// TIA Portal project "e045002v089" (V13) (continued)
VAR_GLOBAL   // PLC tag table "I/O Intercambio Envolvedora"
   "iPalletRetractil" AT %E2.0 : Bool;   // Pallet retractilado (desde el retractilador)
   "oRetractiSeg" AT %A17.7 : Bool;   // Retractilador Seguridades (hacia Retractilador)
   "iPeticionPallet" AT %E2.1 : Bool;   // Petición de pallet (desde el retractilador)
   "oRetractiPermiso" AT %A17.6 : Bool;   // Retractilador Permiso (hacia Retractilador)
   "iBrazoPos_Envolv" AT %E10.5 : Bool;   // Brazo en posición y Freno cerrado en Envolvedora (Retractilador)
   "oHabilMovBrazo_Envol" AT %A16.3 : Bool;   // Habilitación apertura freno brazo Envolvedora (Retractilador)
END_VAR

VAR_GLOBAL   // PLC tag table "I/O Intercambio Cartonero"
   "iCartZonaSeg" AT %M230.1 : Bool;   // Señal de Cartonero: 1= Fuera de zona de paletizadora
   "iCartAplicado" AT %M230.2 : Bool;   // Señal de Cartonero: 1= Cartón aplicado
   "oTomarCartón" AT %A34.3 : Bool;   // Señal a Cartonero: 1= Tomar cartón
   "oAplicarCartón" AT %A34.4 : Bool;   // Señal a Cartonero: 1= Aplicar Cartón
   "oPaleZonaSeg" AT %A34.5 : Bool;   // Señal a Cartonero: 1= Paletizadora en zona segura para el cartonero
   "oPaleSinAlarm" AT %A34.6 : Bool;   // Señal a Cartonero: 1= Paletizadora sin alarmas
   "iCartSinAlarm" AT %M230.0 : Bool;   // Señal de Cartonero: 1= Sin Alarmas
END_VAR

VAR_GLOBAL   // PLC tag table "260_EtiquetadoraYFechadoras"
   "i_FallEnEtiq" AT %I6.6 : Bool;
   "i_FallEnFechadora1" AT %I10.6 : Bool;
   "iSns_PresCajaEmpujador" AT %I11.0 : Bool;
END_VAR

TYPE "Filas_Receta"
   STRUCT
      Bit_1_Elemento : Array [1..10] of Bool;
      Bit_2_Elemento : Array [1..10] of Bool;
   END_STRUCT;
END_TYPE

TYPE "Capas_Receta"
   STRUCT
      Filas : Array [1..6] of "Filas_Receta";
      Usar_Pistón : Bool;
   END_STRUCT;
END_TYPE

TYPE "Elementos HMI"
   STRUCT
      Figura : Byte;
      Estado : Byte;
      Offset_X : Int;
   END_STRUCT;
END_TYPE

TYPE "Filas HMI"
   STRUCT
      Offset_Y : Int;
      Elemento : Array [1 .. 10] of "Elementos HMI";
   END_STRUCT;
END_TYPE

TYPE "Filas_Proceso"
   STRUCT
      Bit_1_Elemento : Array [1 .. 10] of Bool;
      Bit_2_Elemento : Array [1 .. 10] of Bool;
      Actual_Elemento : Array [1 .. 10] of Bool;
   END_STRUCT;
END_TYPE

TYPE "Capas_Proceso"
   STRUCT
      Fila : Array [1 .. 6] of "Filas_Proceso";
      Usar_Pistón : Bool;
   END_STRUCT;
END_TYPE

TYPE "PETICION_CONTROL"
   STRUCT
      cero : Byte;
      PETICION : Byte;
      PARAMETRO : Array [1 .. 3] of Word;
   END_STRUCT;
END_TYPE

TYPE "Recetas"
   STRUCT
      Nombre : Array [1 .. 50] of Char;
      Cant_Capas_Pallet : Byte;
      Cant_Capas_Distintas : Byte;
      Capa : Array [1 .. 10] of "Capas_Receta";
      Vel_Dosificador : Real;
   END_STRUCT;
END_TYPE

DATA_BLOCK "Proceso Dosificador"   // DB2
{ S7_Optimized_Access := 'FALSE' }
VERSION : 0.1
   VAR
      Cant_Cajas : Word;
      Cant_Pallets : Word;
      Capa_Actual : Byte;
      Elemento_Actual : Byte;
      Elemento_Proximo : Byte;
   END_VAR
BEGIN
END_DATA_BLOCK

DATA_BLOCK "DB_Animación"   // DB3
{ S7_Optimized_Access := 'FALSE' }
VERSION : 0.1
   VAR
      Fila : Array [1 .. 6] of "Filas HMI";
      Fila_SEL : Byte;
      Elemento_SEL : Byte;
      Figura_SEL : Byte;
      FechaHora : Date_And_Time;
      Nro_Receta_Edición : Byte;
      Nombre_Receta_Edición : Array [1..50] of Char;
      Capas_X_Pallet_Edición : Byte;
      CapasDistintas_Edición : Byte;
      Capa_Actual_Edición : Byte;
      Usar_Pistón : Bool;
      Vel_Dosificador : Real;
   END_VAR
BEGIN
END_DATA_BLOCK

DATA_BLOCK "HMI"   // DB5
{ S7_Optimized_Access := 'FALSE' }
VERSION : 0.1
   VAR
      Pls_Inc_Elem : Bool;
      Pls_Dec_Elem : Bool;
      Pls_Elem_Der : Bool;
      Pls_Elem_Izq : Bool;
      Pls_Inc_Fila : Bool;
      Pls_Dec_Fila : Bool;
      Pls_Fila_Sup : Bool;
      Pls_Fila_Inf : Bool;
      Pls_New_Fila : Bool;
      Pls_New_Elem : Bool;
      Pls_Kill_Elem : Bool;
      Pls_WR_Receta : Bool;
      Pls_RD_Receta : Bool;
      Pls_CargarReceta : Bool;
      Imagen_Actual : Word;
      Pls_Inc_Receta : Bool;
      Pls_Dec_Receta : Bool;
      Pls_Inc_Capa : Bool;
      Pls_Dec_Capa : Bool;
      "Pls_Elem_+" : Bool;
      "Pls_Elem_-" : Bool;
      Pls_TerminarPallet : Bool;
      Pls_ResetPallets : Bool;
      Pls_ResetCajas : Bool;
      Pls_SalirImagenIni : Bool;
      Pls_RecambioPallet : Bool;
      TP1_a_TP2 : Bool;
      TP2_a_TP3 : Bool;
      TP3_a_TP4 : Bool;
      TP4_a_TP5 : Bool;
      TP5_a_Desc : Bool;
      Pls_Inc_Figura_Sel : Bool;
      Pls_Inc_Capa_Editando : Bool;
      Pls_Dec_Capa_Editando : Bool;
      Pls_MarMan_Ramp1 : Bool;
      Pls_MarMan_Rol1 : Bool;
      Pls_MarMan_Ramp2 : Bool;
      Pls_MarMan_Rol2 : Bool;
      Hab_Cartonero : Bool;
      Cartones_1_o_2 : Bool;
      hab_etiq : Bool;
      hab_fechadora1 : Bool;
      hab_fechadora2 : Bool;
   END_VAR
BEGIN
END_DATA_BLOCK

DATA_BLOCK "flanco"   // DB6
{ S7_Optimized_Access := 'FALSE' }
VERSION : 0.1
   VAR
      "nHMI.Pls_Inc_Elem" : Bool;
      "nHMI.Pls_Dec_Elem" : Bool;
      "nHMI.Pls_Elem_Der" : Bool;
      "nHMI.Pls_Elem_Izq" : Bool;
      "nHMI.Pls_Inc_Fila" : Bool;
      "nHMI.Pls_Dec_Fila" : Bool;
      "nHMI.Pls_Fila_Sup" : Bool;
      "nHMI.Pls_Fila_Inf" : Bool;
      "pHMI.Pls_New_Fila" : Bool;
      "pHMI.Pls_New_Elem" : Bool;
      "pHMI.Pls_Kill_Elem" : Bool;
      "nHMI.Pls_WR_Receta" : Bool;
      "nHMI.Pls_RD_Receta" : Bool;
      pEditando_Recetas : Bool;
      "nHMI.Pls_Inc_Receta" : Bool;
      "nHMI.Pls_Dec_Receta" : Bool;
      "nHMI.Pls_Inc_Capa" : Bool;
      "nHMI.Pls_Dec_Capa" : Bool;
      "nHMI.Pls_Elem_+" : Bool;
      "nHMI.Pls_Elem_-" : Bool;
      "pHMI.Pls_CargarReceta" : Bool;
      piPul_MarCiclo : Bool;
      piPul_HabTransp : Bool;
      piPul_HabDosif : Bool;
      piPul_HabCargPall : Bool;
      piSnsContadEmbal_1 : Bool;
      piSnsContadEmbal_2 : Bool;
      piSnsContadEmbal_3 : Bool;
      niSnsContadEmbal_1 : Bool;
      niSnsContadEmbal_2 : Bool;
      niSnsContadEmbal_3 : Bool;
      "pAUTO/MAN" : Bool;
      "nAUTO/MAN" : Bool;
      piSnsPerEmpCajAde : Bool;
      niSnsPerEmpCajAde : Bool;
      piPul_MultiArr : Bool;
      niPul_MultiArr : Bool;
      piPul_MultiAba : Bool;
      niPul_MultiAba : Bool;
      piPul_MultiAde : Bool;
      niPul_MultiAde : Bool;
      piPul_MultiAtr : Bool;
      niPul_MultiAtr : Bool;
      piPul_Multi_A : Bool;
      niPul_Multi_A : Bool;
      piPul_Multi_B : Bool;
      niPul_Multi_B : Bool;
      niSnsPlataf_Ade : Bool;
      niSnsPlataf_Atr : Bool;
      piSnsPallTrnsp_2 : Bool;
      niSnsPallTrnsp_2 : Bool;
      piSnsPallRetractil : Bool;
      niSnsPallRetractil : Bool;
      piSnsPallTrnsp_4 : Bool;
      niSnsPallTrnsp_4 : Bool;
      piSnsPallTrnsp_5 : Bool;
      niSnsPallTrnsp_5 : Bool;
      piSnsEmpj_Ade_Par : Bool;
      nPALLET_NO_FUERA_ASCENSOR : Bool;
      pRECAMBIO_PALLET : Bool;
      piSnsPallEnAscen : Bool;
      niSnsPallEnAscen : Bool;
      piSnsAltuPlata_Aba : Bool;
      niSnsAltuPlata_Aba : Bool;
      piSnsAltuPlata_Arr : Bool;
      niSnsAltuPlata_Arr : Bool;
      piSnsAscen_Arr : Bool;
      piSnsAscen_Aba_Par : Bool;
      nEditando_Recetas : Bool;
      "pHMI.Pls_RD_Receta" : Bool;
      p3s4_p3s9 : Bool;
      "pHMI.Pls_Inc_Figura_Sel" : Bool;
      "pHMI.Pls_Inc_Capa_Editando" : Bool;
      "pHMI.Pls_Dec_Capa_Editando" : Bool;
      pS_PriElemCapa : Bool;
      nElemento_DESCARGADO : Bool;
   END_VAR
BEGIN
END_DATA_BLOCK

DATA_BLOCK "Constante"   // DB8
{ S7_Optimized_Access := 'FALSE' }
VERSION : 0.1
   VAR
      HMI_Pixel_Offset_X : Int;
      HMI_Pixel_Offset_Y : Int;
      Elemento_SELECCIONADO : Byte;
      Elemento_PRESENTE : Byte;
      Elemento_AUSENTE : Byte;
   END_VAR
BEGIN
END_DATA_BLOCK

DATA_BLOCK "Proceso Empujador"   // DB51
{ S7_Optimized_Access := 'FALSE' }
VERSION : 0.1
   VAR
      Cant_Cajas : DInt;
      Cant_Pallets : DInt;
      Capa_Actual : Byte;
      Elemento_Actual : Byte;
   END_VAR
BEGIN
END_DATA_BLOCK

DATA_BLOCK "PUNTERO_AREA"   // DB55
{ S7_Optimized_Access := 'FALSE' }
VERSION : 0.1
   VAR
      PETICIÓN : "PETICION_CONTROL";
   END_VAR
BEGIN
END_DATA_BLOCK

DATA_BLOCK "Proceso CargaPallet"   // DB89
{ S7_Optimized_Access := 'FALSE' }
VERSION : 0.1
   VAR
      Cant_Cajas : DInt;
      Cant_Pallets : DInt;
      Capa_Actual : Byte;
   END_VAR
BEGIN
END_DATA_BLOCK

DATA_BLOCK "DB_Velocidades"   // DB99
{ S7_Optimized_Access := 'FALSE' }
VERSION : 0.1
   VAR
      Dosif_LímInf_Vel : Real;
      Dosif_Vel_Len : Real;
      Dosif_Vel_Ráp : Real;
      Dosif_LímSup_Vel : Real;
      Empuj_LímInf_Vel : Real;
      Empuj_VelRáp_Ade : Real;
      Empuj_VelLen_Ade : Real;
      Empuj_VelRáp_Atr : Real;
      Empuj_VelLen_Atr : Real;
      Empuj_Vel_Man : Real;
      Empuj_LímSup_Vel : Real;
      Ascens_LímInf_Vel : Real;
      Ascens_VelRáp_Arr : Real;
      Ascens_VelLen_Arr : Real;
      Ascens_VelRáp_Aba : Real;
      Ascens_VelLen_Aba : Real;
      Ascens_Vel_Man : Real;
      Ascens_LímSup_Vel : Real;
   END_VAR
BEGIN
END_DATA_BLOCK

DATA_BLOCK "TIEMPO"   // DB106
{ S7_Optimized_Access := 'FALSE' }
VERSION : 0.1
   VAR
      EMPUJADOR_MED_CAM : Time;
      DOSIF_GIRA_CAJA : Time;
      DOSIF_PROX_CAJA : Time;
      CARGAPALL_BRAZO_PUESTO : Time;
      ESPERA_HH : Time;
      Parada_2s16 : Time;
      Empuja_Caja : Time;
   END_VAR
BEGIN
END_DATA_BLOCK

DATA_BLOCK "PLC a HMI"   // DB119
{ S7_Optimized_Access := 'FALSE' }
VERSION : 0.1
   VAR
      Almacén_Pallets : Bool;
      Elevador : Bool;
      Seg_Elevador : Bool;
      Transp_2 : Bool;
      Transp_3 : Bool;
      Transp_4 : Bool;
      Transp_5 : Bool;
      Descarga : Bool;
      Avance_1_2 : Bool;
      Avance_2_3 : Bool;
      Avance_3_4 : Bool;
      Avance_4_5 : Bool;
      Avance_5_Desc : Bool;
      ETIQUETAR : Bool;
      CICLO_OK : Bool;
      HOME_PISTON : Bool;
      PEDIDO_ENVOLV : Bool;
      ENVOLVER : Bool;
      PALLET_ENVUELTO : Bool;
      TRANSPORTES_Hab : Bool;
      Seg_Entrada_Envol : Bool;
      Seg_Salida_Envol : Bool;
      oTranspPall1 : Bool;
      oTranspPall2 : Bool;
      oTranspPall3 : Bool;
      oTranspPall3Freno : Bool;
      oTranspPall4 : Bool;
      oTranspPall5 : Bool;
      iBrazoPos_Envolv : Bool;
      oHabilMovBrazo_Envol : Bool;
      iCartZonaSeg : Bool;
      iCartAplicado : Bool;
      iCartConAlarm : Bool;
      oTomarCartón : Bool;
      oAplicarCartón : Bool;
      oPaleZonaSeg : Bool;
      oPaleSinAlarm : Bool;
   END_VAR
BEGIN
END_DATA_BLOCK

DATA_BLOCK "Remanente"   // DB173
{ S7_Optimized_Access := 'FALSE' }
VERSION : 0.1
   VAR
      Set_para_2c13 : Bool;
      Mem_Cartón_Aplicado : Bool;
   END_VAR
BEGIN
END_DATA_BLOCK

DATA_BLOCK "DB_Carton_Manual"   // DB175
{ S7_Optimized_Access := 'FALSE' }
VERSION : 0.1
   VAR
      Catoneo_Manual_Hab : Bool;
      CM_FrenoCiclo : Bool;
      CM_OperDetect : Bool;
      FNeg_OperDetect : Bool;
      FPos_ParaFrenCiclo : Bool;
      M_PrimerCapa : Bool;
      F_PrimerCapa : Bool;
   END_VAR
BEGIN
END_DATA_BLOCK

// folder: Alarmas

DATA_BLOCK "DB_ALA_PRE"   // DB56
{ S7_Optimized_Access := 'FALSE' }
VERSION : 0.1
   VAR
      Falla_9 : Bool;
      Falla_10 : Bool;
      Falla_11 : Bool;
      Falla_12 : Bool;
      Falla_13 : Bool;
      Falla_14 : Bool;
      Falla_15 : Bool;
      Falla_16 : Bool;
      Falla_1 : Bool;
      Falla_2 : Bool;
      Falla_3 : Bool;
      Falla_4 : Bool;
      Falla_5 : Bool;
      Falla_6 : Bool;
      Falla_7 : Bool;
      Falla_8 : Bool;
      Falla_25 : Bool;
      Falla_26 : Bool;
      Falla_27 : Bool;
      Falla_28 : Bool;
      Falla_29 : Bool;
      Falla_30 : Bool;
      Falla_31 : Bool;
      Falla_32 : Bool;
      Falla_17 : Bool;
      Falla_18 : Bool;
      Falla_19 : Bool;
      Falla_20 : Bool;
      Falla_21 : Bool;
      Falla_22 : Bool;
      Falla_23 : Bool;
      Falla_24 : Bool;
      Falla_41 : Bool;
      Falla_42 : Bool;
      Falla_43 : Bool;
      Falla_44 : Bool;
      Falla_45 : Bool;
      Falla_46 : Bool;
      Falla_47 : Bool;
      Falla_48 : Bool;
      Falla_33 : Bool;
      Falla_34 : Bool;
      Falla_35 : Bool;
      Falla_36 : Bool;
      Falla_37 : Bool;
      Falla_38 : Bool;
      Falla_39 : Bool;
      Falla_40 : Bool;
      Falla_57 : Bool;
      Falla_58 : Bool;
      Falla_59 : Bool;
      Falla_60 : Bool;
      Falla_61 : Bool;
      Falla_62 : Bool;
      Falla_63 : Bool;
      Falla_64 : Bool;
      Falla_49 : Bool;
      Falla_50 : Bool;
      Falla_51 : Bool;
      Falla_52 : Bool;
      Falla_53 : Bool;
      Falla_54 : Bool;
      Falla_55 : Bool;
      Falla_56 : Bool;
      Falla_73 : Bool;
      Falla_74 : Bool;
      Falla_75 : Bool;
      Falla_76 : Bool;
      Falla_77 : Bool;
      Falla_78 : Bool;
      Falla_79 : Bool;
      Falla_80 : Bool;
      Falla_65 : Bool;
      Falla_66 : Bool;
      Falla_67 : Bool;
      Falla_68 : Bool;
      Falla_69 : Bool;
      Falla_70 : Bool;
      Falla_71 : Bool;
      Falla_72 : Bool;
      Falla_89 : Bool;
      Falla_90 : Bool;
      Falla_91 : Bool;
      Falla_92 : Bool;
      Falla_93 : Bool;
      Falla_94 : Bool;
      Falla_95 : Bool;
      Falla_96 : Bool;
      Falla_81 : Bool;
      Falla_82 : Bool;
      Falla_83 : Bool;
      Falla_84 : Bool;
      Falla_85 : Bool;
      Falla_86 : Bool;
      Falla_87 : Bool;
      Falla_88 : Bool;
      Falla_105 : Bool;
      Falla_106 : Bool;
      Falla_107 : Bool;
      Falla_108 : Bool;
      Falla_109 : Bool;
      Falla_110 : Bool;
      Falla_111 : Bool;
      Falla_112 : Bool;
      Falla_97 : Bool;
      Falla_98 : Bool;
      Falla_99 : Bool;
      Falla_100 : Bool;
      Falla_101 : Bool;
      Falla_102 : Bool;
      Falla_103 : Bool;
      Falla_104 : Bool;
      Falla_121 : Bool;
      Falla_122 : Bool;
      Falla_123 : Bool;
      Falla_124 : Bool;
      Falla_125 : Bool;
      Falla_126 : Bool;
      Falla_127 : Bool;
      Falla_128 : Bool;
      Falla_113 : Bool;
      Falla_114 : Bool;
      Falla_115 : Bool;
      Falla_116 : Bool;
      Falla_117 : Bool;
      Falla_118 : Bool;
      Falla_119 : Bool;
      Falla_120 : Bool;
   END_VAR
BEGIN
END_DATA_BLOCK

DATA_BLOCK "DB_ALA_MEM"   // DB57
{ S7_Optimized_Access := 'FALSE' }
VERSION : 0.1
   VAR
      Alarma_9 : Bool;
      Alarma_10 : Bool;
      Alarma_11 : Bool;
      Alarma_12 : Bool;
      Alarma_13 : Bool;
      Alarma_14 : Bool;
      Alarma_15 : Bool;
      Alarma_16 : Bool;
      Alarma_1 : Bool;
      Alarma_2 : Bool;
      Alarma_3 : Bool;
      Alarma_4 : Bool;
      Alarma_5 : Bool;
      Alarma_6 : Bool;
      Alarma_7 : Bool;
      Alarma_8 : Bool;
      Alarma_25 : Bool;
      Alarma_26 : Bool;
      Alarma_27 : Bool;
      Alarma_28 : Bool;
      Alarma_29 : Bool;
      Alarma_30 : Bool;
      Alarma_31 : Bool;
      Alarma_32 : Bool;
      Alarma_17 : Bool;
      Alarma_18 : Bool;
      Alarma_19 : Bool;
      Alarma_20 : Bool;
      Alarma_21 : Bool;
      Alarma_22 : Bool;
      Alarma_23 : Bool;
      Alarma_24 : Bool;
      Alarma_41 : Bool;
      Alarma_42 : Bool;
      Alarma_43 : Bool;
      Alarma_44 : Bool;
      Alarma_45 : Bool;
      Alarma_46 : Bool;
      Alarma_47 : Bool;
      Alarma_48 : Bool;
      Alarma_33 : Bool;
      Alarma_34 : Bool;
      Alarma_35 : Bool;
      Alarma_36 : Bool;
      Alarma_37 : Bool;
      Alarma_38 : Bool;
      Alarma_39 : Bool;
      Alarma_40 : Bool;
      Alarma_57 : Bool;
      Alarma_58 : Bool;
      Alarma_59 : Bool;
      Alarma_60 : Bool;
      Alarma_61 : Bool;
      Alarma_62 : Bool;
      Alarma_63 : Bool;
      Alarma_64 : Bool;
      Alarma_49 : Bool;
      Alarma_50 : Bool;
      Alarma_51 : Bool;
      Alarma_52 : Bool;
      Alarma_53 : Bool;
      Alarma_54 : Bool;
      Alarma_55 : Bool;
      Alarma_56 : Bool;
      Alarma_73 : Bool;
      Alarma_74 : Bool;
      Alarma_75 : Bool;
      Alarma_76 : Bool;
      Alarma_77 : Bool;
      Alarma_78 : Bool;
      Alarma_79 : Bool;
      Alarma_80 : Bool;
      Alarma_65 : Bool;
      Alarma_66 : Bool;
      Alarma_67 : Bool;
      Alarma_68 : Bool;
      Alarma_69 : Bool;
      Alarma_70 : Bool;
      Alarma_71 : Bool;
      Alarma_72 : Bool;
      Alarma_89 : Bool;
      Alarma_90 : Bool;
      Alarma_91 : Bool;
      Alarma_92 : Bool;
      Alarma_93 : Bool;
      Alarma_94 : Bool;
      Alarma_95 : Bool;
      Alarma_96 : Bool;
      Alarma_81 : Bool;
      Alarma_82 : Bool;
      Alarma_83 : Bool;
      Alarma_84 : Bool;
      Alarma_85 : Bool;
      Alarma_86 : Bool;
      Alarma_87 : Bool;
      Alarma_88 : Bool;
      Alarma_105 : Bool;
      Alarma_106 : Bool;
      Alarma_107 : Bool;
      Alarma_108 : Bool;
      Alarma_109 : Bool;
      Alarma_110 : Bool;
      Alarma_111 : Bool;
      Alarma_112 : Bool;
      Alarma_97 : Bool;
      Alarma_98 : Bool;
      Alarma_99 : Bool;
      Alarma_100 : Bool;
      Alarma_101 : Bool;
      Alarma_102 : Bool;
      Alarma_103 : Bool;
      Alarma_104 : Bool;
      Alarma_121 : Bool;
      Alarma_122 : Bool;
      Alarma_123 : Bool;
      Alarma_124 : Bool;
      Alarma_125 : Bool;
      Alarma_126 : Bool;
      Alarma_127 : Bool;
      Alarma_128 : Bool;
      Alarma_113 : Bool;
      Alarma_114 : Bool;
      Alarma_115 : Bool;
      Alarma_116 : Bool;
      Alarma_117 : Bool;
      Alarma_118 : Bool;
      Alarma_119 : Bool;
      Alarma_120 : Bool;
   END_VAR
BEGIN
END_DATA_BLOCK

DATA_BLOCK "DB_ALA_REC"   // DB58
{ S7_Optimized_Access := 'FALSE' }
VERSION : 0.1
   VAR
      AlaRec_9 : Bool;
      AlaRec_10 : Bool;
      AlaRec_11 : Bool;
      AlaRec_12 : Bool;
      AlaRec_13 : Bool;
      AlaRec_14 : Bool;
      AlaRec_15 : Bool;
      AlaRec_16 : Bool;
      AlaRec_1 : Bool;
      AlaRec_2 : Bool;
      AlaRec_3 : Bool;
      AlaRec_4 : Bool;
      AlaRec_5 : Bool;
      AlaRec_6 : Bool;
      AlaRec_7 : Bool;
      AlaRec_8 : Bool;
      AlaRec_25 : Bool;
      AlaRec_26 : Bool;
      AlaRec_27 : Bool;
      AlaRec_28 : Bool;
      AlaRec_29 : Bool;
      AlaRec_30 : Bool;
      AlaRec_31 : Bool;
      AlaRec_32 : Bool;
      AlaRec_17 : Bool;
      AlaRec_18 : Bool;
      AlaRec_19 : Bool;
      AlaRec_20 : Bool;
      AlaRec_21 : Bool;
      AlaRec_22 : Bool;
      AlaRec_23 : Bool;
      AlaRec_24 : Bool;
      AlaRec_41 : Bool;
      AlaRec_42 : Bool;
      AlaRec_43 : Bool;
      AlaRec_44 : Bool;
      AlaRec_45 : Bool;
      AlaRec_46 : Bool;
      AlaRec_47 : Bool;
      AlaRec_48 : Bool;
      AlaRec_33 : Bool;
      AlaRec_34 : Bool;
      AlaRec_35 : Bool;
      AlaRec_36 : Bool;
      AlaRec_37 : Bool;
      AlaRec_38 : Bool;
      AlaRec_39 : Bool;
      AlaRec_40 : Bool;
      AlaRec_57 : Bool;
      AlaRec_58 : Bool;
      AlaRec_59 : Bool;
      AlaRec_60 : Bool;
      AlaRec_61 : Bool;
      AlaRec_62 : Bool;
      AlaRec_63 : Bool;
      AlaRec_64 : Bool;
      AlaRec_49 : Bool;
      AlaRec_50 : Bool;
      AlaRec_51 : Bool;
      AlaRec_52 : Bool;
      AlaRec_53 : Bool;
      AlaRec_54 : Bool;
      AlaRec_55 : Bool;
      AlaRec_56 : Bool;
      AlaRec_73 : Bool;
      AlaRec_74 : Bool;
      AlaRec_75 : Bool;
      AlaRec_76 : Bool;
      AlaRec_77 : Bool;
      AlaRec_78 : Bool;
      AlaRec_79 : Bool;
      AlaRec_80 : Bool;
      AlaRec_65 : Bool;
      AlaRec_66 : Bool;
      AlaRec_67 : Bool;
      AlaRec_68 : Bool;
      AlaRec_69 : Bool;
      AlaRec_70 : Bool;
      AlaRec_71 : Bool;
      AlaRec_72 : Bool;
      AlaRec_89 : Bool;
      AlaRec_90 : Bool;
      AlaRec_91 : Bool;
      AlaRec_92 : Bool;
      AlaRec_93 : Bool;
      AlaRec_94 : Bool;
      AlaRec_95 : Bool;
      AlaRec_96 : Bool;
      AlaRec_81 : Bool;
      AlaRec_82 : Bool;
      AlaRec_83 : Bool;
      AlaRec_84 : Bool;
      AlaRec_85 : Bool;
      AlaRec_86 : Bool;
      AlaRec_87 : Bool;
      AlaRec_88 : Bool;
      AlaRec_105 : Bool;
      AlaRec_106 : Bool;
      AlaRec_107 : Bool;
      AlaRec_108 : Bool;
      AlaRec_109 : Bool;
      AlaRec_110 : Bool;
      AlaRec_111 : Bool;
      AlaRec_112 : Bool;
      AlaRec_97 : Bool;
      AlaRec_98 : Bool;
      AlaRec_99 : Bool;
      AlaRec_100 : Bool;
      AlaRec_101 : Bool;
      AlaRec_102 : Bool;
      AlaRec_103 : Bool;
      AlaRec_104 : Bool;
      AlaRec_121 : Bool;
      AlaRec_122 : Bool;
      AlaRec_123 : Bool;
      AlaRec_124 : Bool;
      AlaRec_125 : Bool;
      AlaRec_126 : Bool;
      AlaRec_127 : Bool;
      AlaRec_128 : Bool;
      AlaRec_113 : Bool;
      AlaRec_114 : Bool;
      AlaRec_115 : Bool;
      AlaRec_116 : Bool;
      AlaRec_117 : Bool;
      AlaRec_118 : Bool;
      AlaRec_119 : Bool;
      AlaRec_120 : Bool;
   END_VAR
BEGIN
END_DATA_BLOCK

DATA_BLOCK "DB_COM_REC"   // DB59
{ S7_Optimized_Access := 'FALSE' }
VERSION : 0.1
   VAR
      ComRec_9 : Bool;
      ComRec_10 : Bool;
      ComRec_11 : Bool;
      ComRec_12 : Bool;
      ComRec_13 : Bool;
      ComRec_14 : Bool;
      ComRec_15 : Bool;
      ComRec_16 : Bool;
      ComRec_1 : Bool;
      ComRec_2 : Bool;
      ComRec_3 : Bool;
      ComRec_4 : Bool;
      ComRec_5 : Bool;
      ComRec_6 : Bool;
      ComRec_7 : Bool;
      ComRec_8 : Bool;
      ComRec_25 : Bool;
      ComRec_26 : Bool;
      ComRec_27 : Bool;
      ComRec_28 : Bool;
      ComRec_29 : Bool;
      ComRec_30 : Bool;
      ComRec_31 : Bool;
      ComRec_32 : Bool;
      ComRec_17 : Bool;
      ComRec_18 : Bool;
      ComRec_19 : Bool;
      ComRec_20 : Bool;
      ComRec_21 : Bool;
      ComRec_22 : Bool;
      ComRec_23 : Bool;
      ComRec_24 : Bool;
      ComRec_41 : Bool;
      ComRec_42 : Bool;
      ComRec_43 : Bool;
      ComRec_44 : Bool;
      ComRec_45 : Bool;
      ComRec_46 : Bool;
      ComRec_47 : Bool;
      ComRec_48 : Bool;
      ComRec_33 : Bool;
      ComRec_34 : Bool;
      ComRec_35 : Bool;
      ComRec_36 : Bool;
      ComRec_37 : Bool;
      ComRec_38 : Bool;
      ComRec_39 : Bool;
      ComRec_40 : Bool;
      ComRec_57 : Bool;
      ComRec_58 : Bool;
      ComRec_59 : Bool;
      ComRec_60 : Bool;
      ComRec_61 : Bool;
      ComRec_62 : Bool;
      ComRec_63 : Bool;
      ComRec_64 : Bool;
      ComRec_49 : Bool;
      ComRec_50 : Bool;
      ComRec_51 : Bool;
      ComRec_52 : Bool;
      ComRec_53 : Bool;
      ComRec_54 : Bool;
      ComRec_55 : Bool;
      ComRec_56 : Bool;
      ComRec_73 : Bool;
      ComRec_74 : Bool;
      ComRec_75 : Bool;
      ComRec_76 : Bool;
      ComRec_77 : Bool;
      ComRec_78 : Bool;
      ComRec_79 : Bool;
      ComRec_80 : Bool;
      ComRec_65 : Bool;
      ComRec_66 : Bool;
      ComRec_67 : Bool;
      ComRec_68 : Bool;
      ComRec_69 : Bool;
      ComRec_70 : Bool;
      ComRec_71 : Bool;
      ComRec_72 : Bool;
      ComRec_89 : Bool;
      ComRec_90 : Bool;
      ComRec_91 : Bool;
      ComRec_92 : Bool;
      ComRec_93 : Bool;
      ComRec_94 : Bool;
      ComRec_95 : Bool;
      ComRec_96 : Bool;
      ComRec_81 : Bool;
      ComRec_82 : Bool;
      ComRec_83 : Bool;
      ComRec_84 : Bool;
      ComRec_85 : Bool;
      ComRec_86 : Bool;
      ComRec_87 : Bool;
      ComRec_88 : Bool;
      ComRec_105 : Bool;
      ComRec_106 : Bool;
      ComRec_107 : Bool;
      ComRec_108 : Bool;
      ComRec_109 : Bool;
      ComRec_110 : Bool;
      ComRec_111 : Bool;
      ComRec_112 : Bool;
      ComRec_97 : Bool;
      ComRec_98 : Bool;
      ComRec_99 : Bool;
      ComRec_100 : Bool;
      ComRec_101 : Bool;
      ComRec_102 : Bool;
      ComRec_103 : Bool;
      ComRec_104 : Bool;
      ComRec_121 : Bool;
      ComRec_122 : Bool;
      ComRec_123 : Bool;
      ComRec_124 : Bool;
      ComRec_125 : Bool;
      ComRec_126 : Bool;
      ComRec_127 : Bool;
      ComRec_128 : Bool;
      ComRec_113 : Bool;
      ComRec_114 : Bool;
      ComRec_115 : Bool;
      ComRec_116 : Bool;
      ComRec_117 : Bool;
      ComRec_118 : Bool;
      ComRec_119 : Bool;
      ComRec_120 : Bool;
   END_VAR
BEGIN
END_DATA_BLOCK

DATA_BLOCK "DB_COM_REC_FLANCO"   // DB60
{ S7_Optimized_Access := 'FALSE' }
VERSION : 0.1
   VAR
      ComRecFlanco_9 : Bool;
      ComRecFlanco_10 : Bool;
      ComRecFlanco_11 : Bool;
      ComRecFlanco_12 : Bool;
      ComRecFlanco_13 : Bool;
      ComRecFlanco_14 : Bool;
      ComRecFlanco_15 : Bool;
      ComRecFlanco_16 : Bool;
      ComRecFlanco_1 : Bool;
      ComRecFlanco_2 : Bool;
      ComRecFlanco_3 : Bool;
      ComRecFlanco_4 : Bool;
      ComRecFlanco_5 : Bool;
      ComRecFlanco_6 : Bool;
      ComRecFlanco_7 : Bool;
      ComRecFlanco_8 : Bool;
      ComRecFlanco_25 : Bool;
      ComRecFlanco_26 : Bool;
      ComRecFlanco_27 : Bool;
      ComRecFlanco_28 : Bool;
      ComRecFlanco_29 : Bool;
      ComRecFlanco_30 : Bool;
      ComRecFlanco_31 : Bool;
      ComRecFlanco_32 : Bool;
      ComRecFlanco_17 : Bool;
      ComRecFlanco_18 : Bool;
      ComRecFlanco_19 : Bool;
      ComRecFlanco_20 : Bool;
      ComRecFlanco_21 : Bool;
      ComRecFlanco_22 : Bool;
      ComRecFlanco_23 : Bool;
      ComRecFlanco_24 : Bool;
      ComRecFlanco_41 : Bool;
      ComRecFlanco_42 : Bool;
      ComRecFlanco_43 : Bool;
      ComRecFlanco_44 : Bool;
      ComRecFlanco_45 : Bool;
      ComRecFlanco_46 : Bool;
      ComRecFlanco_47 : Bool;
      ComRecFlanco_48 : Bool;
      ComRecFlanco_33 : Bool;
      ComRecFlanco_34 : Bool;
      ComRecFlanco_35 : Bool;
      ComRecFlanco_36 : Bool;
      ComRecFlanco_37 : Bool;
      ComRecFlanco_38 : Bool;
      ComRecFlanco_39 : Bool;
      ComRecFlanco_40 : Bool;
      ComRecFlanco_57 : Bool;
      ComRecFlanco_58 : Bool;
      ComRecFlanco_59 : Bool;
      ComRecFlanco_60 : Bool;
      ComRecFlanco_61 : Bool;
      ComRecFlanco_62 : Bool;
      ComRecFlanco_63 : Bool;
      ComRecFlanco_64 : Bool;
      ComRecFlanco_49 : Bool;
      ComRecFlanco_50 : Bool;
      ComRecFlanco_51 : Bool;
      ComRecFlanco_52 : Bool;
      ComRecFlanco_53 : Bool;
      ComRecFlanco_54 : Bool;
      ComRecFlanco_55 : Bool;
      ComRecFlanco_56 : Bool;
      ComRecFlanco_73 : Bool;
      ComRecFlanco_74 : Bool;
      ComRecFlanco_75 : Bool;
      ComRecFlanco_76 : Bool;
      ComRecFlanco_77 : Bool;
      ComRecFlanco_78 : Bool;
      ComRecFlanco_79 : Bool;
      ComRecFlanco_80 : Bool;
      ComRecFlanco_65 : Bool;
      ComRecFlanco_66 : Bool;
      ComRecFlanco_67 : Bool;
      ComRecFlanco_68 : Bool;
      ComRecFlanco_69 : Bool;
      ComRecFlanco_70 : Bool;
      ComRecFlanco_71 : Bool;
      ComRecFlanco_72 : Bool;
      ComRecFlanco_89 : Bool;
      ComRecFlanco_90 : Bool;
      ComRecFlanco_91 : Bool;
      ComRecFlanco_92 : Bool;
      ComRecFlanco_93 : Bool;
      ComRecFlanco_94 : Bool;
      ComRecFlanco_95 : Bool;
      ComRecFlanco_96 : Bool;
      ComRecFlanco_81 : Bool;
      ComRecFlanco_82 : Bool;
      ComRecFlanco_83 : Bool;
      ComRecFlanco_84 : Bool;
      ComRecFlanco_85 : Bool;
      ComRecFlanco_86 : Bool;
      ComRecFlanco_87 : Bool;
      ComRecFlanco_88 : Bool;
      ComRecFlanco_105 : Bool;
      ComRecFlanco_106 : Bool;
      ComRecFlanco_107 : Bool;
      ComRecFlanco_108 : Bool;
      ComRecFlanco_109 : Bool;
      ComRecFlanco_110 : Bool;
      ComRecFlanco_111 : Bool;
      ComRecFlanco_112 : Bool;
      ComRecFlanco_97 : Bool;
      ComRecFlanco_98 : Bool;
      ComRecFlanco_99 : Bool;
      ComRecFlanco_100 : Bool;
      ComRecFlanco_101 : Bool;
      ComRecFlanco_102 : Bool;
      ComRecFlanco_103 : Bool;
      ComRecFlanco_104 : Bool;
      ComRecFlanco_121 : Bool;
      ComRecFlanco_122 : Bool;
      ComRecFlanco_123 : Bool;
      ComRecFlanco_124 : Bool;
      ComRecFlanco_125 : Bool;
      ComRecFlanco_126 : Bool;
      ComRecFlanco_127 : Bool;
      ComRecFlanco_128 : Bool;
      ComRecFlanco_113 : Bool;
      ComRecFlanco_114 : Bool;
      ComRecFlanco_115 : Bool;
      ComRecFlanco_116 : Bool;
      ComRecFlanco_117 : Bool;
      ComRecFlanco_118 : Bool;
      ComRecFlanco_119 : Bool;
      ComRecFlanco_120 : Bool;
   END_VAR
BEGIN
END_DATA_BLOCK

DATA_BLOCK "DB_COM_REC_AUX"   // DB61
{ S7_Optimized_Access := 'FALSE' }
VERSION : 0.1
   VAR
      ComRecAux_9 : Bool;
      ComRecAux_10 : Bool;
      ComRecAux_11 : Bool;
      ComRecAux_12 : Bool;
      ComRecAux_13 : Bool;
      ComRecAux_14 : Bool;
      ComRecAux_15 : Bool;
      ComRecAux_16 : Bool;
      ComRecAux_1 : Bool;
      ComRecAux_2 : Bool;
      ComRecAux_3 : Bool;
      ComRecAux_4 : Bool;
      ComRecAux_5 : Bool;
      ComRecAux_6 : Bool;
      ComRecAux_7 : Bool;
      ComRecAux_8 : Bool;
      ComRecAux_25 : Bool;
      ComRecAux_26 : Bool;
      ComRecAux_27 : Bool;
      ComRecAux_28 : Bool;
      ComRecAux_29 : Bool;
      ComRecAux_30 : Bool;
      ComRecAux_31 : Bool;
      ComRecAux_32 : Bool;
      ComRecAux_17 : Bool;
      ComRecAux_18 : Bool;
      ComRecAux_19 : Bool;
      ComRecAux_20 : Bool;
      ComRecAux_21 : Bool;
      ComRecAux_22 : Bool;
      ComRecAux_23 : Bool;
      ComRecAux_24 : Bool;
      ComRecAux_41 : Bool;
      ComRecAux_42 : Bool;
      ComRecAux_43 : Bool;
      ComRecAux_44 : Bool;
      ComRecAux_45 : Bool;
      ComRecAux_46 : Bool;
      ComRecAux_47 : Bool;
      ComRecAux_48 : Bool;
      ComRecAux_33 : Bool;
      ComRecAux_34 : Bool;
      ComRecAux_35 : Bool;
      ComRecAux_36 : Bool;
      ComRecAux_37 : Bool;
      ComRecAux_38 : Bool;
      ComRecAux_39 : Bool;
      ComRecAux_40 : Bool;
      ComRecAux_57 : Bool;
      ComRecAux_58 : Bool;
      ComRecAux_59 : Bool;
      ComRecAux_60 : Bool;
      ComRecAux_61 : Bool;
      ComRecAux_62 : Bool;
      ComRecAux_63 : Bool;
      ComRecAux_64 : Bool;
      ComRecAux_49 : Bool;
      ComRecAux_50 : Bool;
      ComRecAux_51 : Bool;
      ComRecAux_52 : Bool;
      ComRecAux_53 : Bool;
      ComRecAux_54 : Bool;
      ComRecAux_55 : Bool;
      ComRecAux_56 : Bool;
      ComRecAux_73 : Bool;
      ComRecAux_74 : Bool;
      ComRecAux_75 : Bool;
      ComRecAux_76 : Bool;
      ComRecAux_77 : Bool;
      ComRecAux_78 : Bool;
      ComRecAux_79 : Bool;
      ComRecAux_80 : Bool;
      ComRecAux_65 : Bool;
      ComRecAux_66 : Bool;
      ComRecAux_67 : Bool;
      ComRecAux_68 : Bool;
      ComRecAux_69 : Bool;
      ComRecAux_70 : Bool;
      ComRecAux_71 : Bool;
      ComRecAux_72 : Bool;
      ComRecAux_89 : Bool;
      ComRecAux_90 : Bool;
      ComRecAux_91 : Bool;
      ComRecAux_92 : Bool;
      ComRecAux_93 : Bool;
      ComRecAux_94 : Bool;
      ComRecAux_95 : Bool;
      ComRecAux_96 : Bool;
      ComRecAux_81 : Bool;
      ComRecAux_82 : Bool;
      ComRecAux_83 : Bool;
      ComRecAux_84 : Bool;
      ComRecAux_85 : Bool;
      ComRecAux_86 : Bool;
      ComRecAux_87 : Bool;
      ComRecAux_88 : Bool;
      ComRecAux_105 : Bool;
      ComRecAux_106 : Bool;
      ComRecAux_107 : Bool;
      ComRecAux_108 : Bool;
      ComRecAux_109 : Bool;
      ComRecAux_110 : Bool;
      ComRecAux_111 : Bool;
      ComRecAux_112 : Bool;
      ComRecAux_97 : Bool;
      ComRecAux_98 : Bool;
      ComRecAux_99 : Bool;
      ComRecAux_100 : Bool;
      ComRecAux_101 : Bool;
      ComRecAux_102 : Bool;
      ComRecAux_103 : Bool;
      ComRecAux_104 : Bool;
      ComRecAux_121 : Bool;
      ComRecAux_122 : Bool;
      ComRecAux_123 : Bool;
      ComRecAux_124 : Bool;
      ComRecAux_125 : Bool;
      ComRecAux_126 : Bool;
      ComRecAux_127 : Bool;
      ComRecAux_128 : Bool;
      ComRecAux_113 : Bool;
      ComRecAux_114 : Bool;
      ComRecAux_115 : Bool;
      ComRecAux_116 : Bool;
      ComRecAux_117 : Bool;
      ComRecAux_118 : Bool;
      ComRecAux_119 : Bool;
      ComRecAux_120 : Bool;
   END_VAR
BEGIN
END_DATA_BLOCK

DATA_BLOCK "DB_BIT_VIDA"   // DB62
{ S7_Optimized_Access := 'FALSE' }
VERSION : 0.1
   VAR
      BitVida_9 : Bool;
      BitVida_10 : Bool;
      BitVida_11 : Bool;
      BitVida_12 : Bool;
      BitVida_13 : Bool;
      BitVida_14 : Bool;
      BitVida_15 : Bool;
      BitVida_16 : Bool;
      BitVida_1 : Bool;
      BitVida_2 : Bool;
      BitVida_3 : Bool;
      BitVida_4 : Bool;
      BitVida_5 : Bool;
      BitVida_6 : Bool;
      BitVida_7 : Bool;
      BitVida_8 : Bool;
      BitVida_25 : Bool;
      BitVida_26 : Bool;
      BitVida_27 : Bool;
      BitVida_28 : Bool;
      BitVida_29 : Bool;
      BitVida_30 : Bool;
      BitVida_31 : Bool;
      BitVida_32 : Bool;
      BitVida_17 : Bool;
      BitVida_18 : Bool;
      BitVida_19 : Bool;
      BitVida_20 : Bool;
      BitVida_21 : Bool;
      BitVida_22 : Bool;
      BitVida_23 : Bool;
      BitVida_24 : Bool;
      BitVida_41 : Bool;
      BitVida_42 : Bool;
      BitVida_43 : Bool;
      BitVida_44 : Bool;
      BitVida_45 : Bool;
      BitVida_46 : Bool;
      BitVida_47 : Bool;
      BitVida_48 : Bool;
      BitVida_33 : Bool;
      BitVida_34 : Bool;
      BitVida_35 : Bool;
      BitVida_36 : Bool;
      BitVida_37 : Bool;
      BitVida_38 : Bool;
      BitVida_39 : Bool;
      BitVida_40 : Bool;
      BitVida_57 : Bool;
      BitVida_58 : Bool;
      BitVida_59 : Bool;
      BitVida_60 : Bool;
      BitVida_61 : Bool;
      BitVida_62 : Bool;
      BitVida_63 : Bool;
      BitVida_64 : Bool;
      BitVida_49 : Bool;
      BitVida_50 : Bool;
      BitVida_51 : Bool;
      BitVida_52 : Bool;
      BitVida_53 : Bool;
      BitVida_54 : Bool;
      BitVida_55 : Bool;
      BitVida_56 : Bool;
      BitVida_73 : Bool;
      BitVida_74 : Bool;
      BitVida_75 : Bool;
      BitVida_76 : Bool;
      BitVida_77 : Bool;
      BitVida_78 : Bool;
      BitVida_79 : Bool;
      BitVida_80 : Bool;
      BitVida_65 : Bool;
      BitVida_66 : Bool;
      BitVida_67 : Bool;
      BitVida_68 : Bool;
      BitVida_69 : Bool;
      BitVida_70 : Bool;
      BitVida_71 : Bool;
      BitVida_72 : Bool;
      BitVida_89 : Bool;
      BitVida_90 : Bool;
      BitVida_91 : Bool;
      BitVida_92 : Bool;
      BitVida_93 : Bool;
      BitVida_94 : Bool;
      BitVida_95 : Bool;
      BitVida_96 : Bool;
      BitVida_81 : Bool;
      BitVida_82 : Bool;
      BitVida_83 : Bool;
      BitVida_84 : Bool;
      BitVida_85 : Bool;
      BitVida_86 : Bool;
      BitVida_87 : Bool;
      BitVida_88 : Bool;
      BitVida_105 : Bool;
      BitVida_106 : Bool;
      BitVida_107 : Bool;
      BitVida_108 : Bool;
      BitVida_109 : Bool;
      BitVida_110 : Bool;
      BitVida_111 : Bool;
      BitVida_112 : Bool;
      BitVida_97 : Bool;
      BitVida_98 : Bool;
      BitVida_99 : Bool;
      BitVida_100 : Bool;
      BitVida_101 : Bool;
      BitVida_102 : Bool;
      BitVida_103 : Bool;
      BitVida_104 : Bool;
      BitVida_121 : Bool;
      BitVida_122 : Bool;
      BitVida_123 : Bool;
      BitVida_124 : Bool;
      BitVida_125 : Bool;
      BitVida_126 : Bool;
      BitVida_127 : Bool;
      BitVida_128 : Bool;
      BitVida_113 : Bool;
      BitVida_114 : Bool;
      BitVida_115 : Bool;
      BitVida_116 : Bool;
      BitVida_117 : Bool;
      BitVida_118 : Bool;
      BitVida_119 : Bool;
      BitVida_120 : Bool;
   END_VAR
BEGIN
END_DATA_BLOCK

// folder: Instancias

DATA_BLOCK "VARIADOR_DOSIFICADOR"   // DB15
{ S7_Optimized_Access := 'FALSE' }
VERSION : 0.1
// stored: InstanceOfName FB_VAR_MOT
"FB_VAR_MOT"
BEGIN
END_DATA_BLOCK

DATA_BLOCK "GIRA_CAJA"   // DB18
{ S7_Optimized_Access := 'FALSE' }
VERSION : 0.1
// stored: InstanceOfName FB_CTR_VAL
"FB_CTR_VAL"
BEGIN
END_DATA_BLOCK

DATA_BLOCK "EMPUJA_CAJA"   // DB19
{ S7_Optimized_Access := 'FALSE' }
VERSION : 0.1
// stored: InstanceOfName FB_CTR_VAL
"FB_CTR_VAL"
BEGIN
END_DATA_BLOCK

DATA_BLOCK "STOP_CAJA"   // DB20
{ S7_Optimized_Access := 'FALSE' }
VERSION : 0.1
// stored: InstanceOfName FB_CTR_VAL
"FB_CTR_VAL"
BEGIN
END_DATA_BLOCK

DATA_BLOCK "VARIADOR_ASCENSOR"   // DB36
{ S7_Optimized_Access := 'FALSE' }
VERSION : 0.1
// stored: InstanceOfName FB_VAR_MOT
"FB_VAR_MOT"
BEGIN
END_DATA_BLOCK

DATA_BLOCK "BRAZO_PLATAFORMA"   // DB37
{ S7_Optimized_Access := 'FALSE' }
VERSION : 0.1
// stored: InstanceOfName FB_CTR_VAL
"FB_CTR_VAL"
BEGIN
END_DATA_BLOCK

DATA_BLOCK "EMPUJADOR_EN_BRAZO"   // DB38
{ S7_Optimized_Access := 'FALSE' }
VERSION : 0.1
// stored: InstanceOfName FB_CTR_VAL
"FB_CTR_VAL"
BEGIN
END_DATA_BLOCK

DATA_BLOCK "MORDAZAS_LATERALES"   // DB39
{ S7_Optimized_Access := 'FALSE' }
VERSION : 0.1
// stored: InstanceOfName FB_CTR_VAL
"FB_CTR_VAL"
BEGIN
END_DATA_BLOCK

DATA_BLOCK "MORDAZA_FINAL"   // DB40
{ S7_Optimized_Access := 'FALSE' }
VERSION : 0.1
// stored: InstanceOfName FB_CTR_VAL
"FB_CTR_VAL"
BEGIN
END_DATA_BLOCK

DATA_BLOCK "EMPUJADOR_FILAS_ADELANTE/ATRÁS"   // DB53
{ S7_Optimized_Access := 'FALSE' }
VERSION : 0.1
// stored: InstanceOfName FB_VAR_MOT
"FB_VAR_MOT"
BEGIN
END_DATA_BLOCK

DATA_BLOCK "ALMACÉN_PALLET"   // DB69
{ S7_Optimized_Access := 'FALSE' }
VERSION : 0.1
// stored: InstanceOfName FB_CTR_VAL
"FB_CTR_VAL"
BEGIN
END_DATA_BLOCK

DATA_BLOCK "DEDOS_ALMACÉN"   // DB70
{ S7_Optimized_Access := 'FALSE' }
VERSION : 0.1
// stored: InstanceOfName FB_CTR_VAL
"FB_CTR_VAL"
BEGIN
END_DATA_BLOCK